
   "Z201".tInputs.xM209FanProtection :="FB_CommunicationZ300_V1.00_DB".IN_tIDeviceDataIN.Z200.IN_MCC1201."xA.E83.5";
   "Z201".tInputs.xM209FanFeedback := "FB_CommunicationZ300_V1.00_DB".IN_tIDeviceDataIN.Z200.IN_MCC1201."xA.E83.6";

   "FB_ManInsp_V1_00_IDB".INPUT.rgxQualityButtons[1]:="FB_CommunicationZ300_V1.00_DB".IN_tIDeviceDataIN.Z200.IN_MCC1301."xE.E108.4";


   "FB_DropConveyor_IDB".INPUT.xUpPosition := "FB_CommunicationZ300_V1.00_DB".IN_tIDeviceDataIN.Z200.IN_MCC1201."xA.E82.1";
   "FB_DropConveyor_IDB".INPUT.xDownPosition := "FB_CommunicationZ300_V1.00_DB".IN_tIDeviceDataIN.Z200.IN_MCC1201."xA.E82.2";
   "FB_DropConveyor_IDB".INPUT.xDoorOpen := "FB_CommunicationZ300_V1.00_DB".IN_tIDeviceDataIN.Z200.IN_MCC1201."xA.E34.0"OR"FB_CommunicationZ300_V1.00_DB".IN_tIDeviceDataIN.Z200.IN_MCC1201."xA.E34.7" ;
   "FB_DropConveyor_IDB".INPUT.xFeedbackMovement :="FB_CommunicationZ300_V1.00_DB".IN_tIDeviceDataIN.Z200.IN_MCC1201."xA.E82.0" ;
   "FB_DropConveyor_IDB".INPUT.xProtection :="FB_CommunicationZ300_V1.00_DB".IN_tIDeviceDataIN.Z200.IN_MCC1201."xA.E81.5" ;
   "FB_DropConveyor_IDB".INPUT.xProtectionBrake := 1;
   "FB_DropConveyor_IDB".INPUT.xUpDownPushbutton := "FB_CommunicationZ300_V1.00_DB".IN_tIDeviceDataIN.Z200.IN_MCC1201."xA.E35.0" OR"FB_CommunicationZ300_V1.00_DB".IN_tIDeviceDataIN.Z200.IN_MCC1201."xA.E34.2" ;
   "FB_DropConveyor_IDB".INPUT.xSafetyBar := "FB_CommunicationZ300_V1.00_DB".IN_tIDeviceDataIN.Z200.IN_MCC1201."xA.E82.3";

   "FB_BreakerM206_V1_00_IDB".INPUT.xConditionOKFromCulletSystem := "FB_CommunicationZ300_V1.00_DB".IN_tIDeviceDataIN.Z200.IN_MCC1201."xA.E39.0";
   "FB_BreakerM206_V1_00_IDB".INPUT.xBreakerRotationControl := "FB_CommunicationZ300_V1.00_DB".IN_tIDeviceDataIN.Z200.IN_MCC1201."xA.E36.0";
   "FB_BreakerM206_V1_00_IDB".INPUT.xProtectionBreakerRotation := "FB_CommunicationZ300_V1.00_DB".IN_tIDeviceDataIN.Z200.IN_MCC1201."xA.E83.0";
   "FB_BreakerM206_V1_00_IDB".INPUT.xFeedbackRotationKM := "FB_CommunicationZ300_V1.00_DB".IN_tIDeviceDataIN.Z200.IN_MCC1201."xA.E83.1";

   "FB_IO_EmergencyCuttingBridge_DB".IN_xMachineReady :="FB_CommunicationZ300_V1.00_DB".IN_tIDeviceDataIN.Z200.IN_MCC1201."xA.E33.4";
   "FB_IO_EmergencyCuttingBridge_DB".IN_xStartCutCycle := "FB_CommunicationZ300_V1.00_DB".IN_tIDeviceDataIN.Z200.IN_MCC1201."xA.E33.5";
   "FB_IO_EmergencyCuttingBridge_DB".IN_xProtection := "FB_CommunicationZ300_V1.00_DB".IN_tIDeviceDataIN.Z200.IN_MCC1201."xA.E81.2";

   "FB_BD_BreakPH_V1_00_IDB".INPUT.rgxPhotoStatus[0] := "FB_CommunicationZ300_V1.00_DB".IN_tIDeviceDataIN.Z200.IN_MCC1201."xA.E32.0";
   "FB_BD_BreakPH_V1_00_IDB".INPUT.rgxPhotoStatus[1]:= "FB_CommunicationZ300_V1.00_DB".IN_tIDeviceDataIN.Z200.IN_MCC1201."xA.E32.1";
   "FB_BD_BreakPH_V1_00_IDB".INPUT.rgxPhotoStatus[2] := "FB_CommunicationZ300_V1.00_DB".IN_tIDeviceDataIN.Z200.IN_MCC1201."xA.E32.2";
   "FB_BD_BreakPH_V1_00_IDB".INPUT.rgxPhotoStatus[3] := "FB_CommunicationZ300_V1.00_DB".IN_tIDeviceDataIN.Z200.IN_MCC1201."xA.E32.3";
   "FB_BD_BreakPH_V1_00_IDB".INPUT.rgxPhotoStatus[4] := "FB_CommunicationZ300_V1.00_DB".IN_tIDeviceDataIN.Z200.IN_MCC1201."xA.E32.4";
   "FB_BD_BreakPH_V1_00_IDB".INPUT.rgxPhotoStatus[5] := "FB_CommunicationZ300_V1.00_DB".IN_tIDeviceDataIN.Z200.IN_MCC1201."xA.E32.5";
   "FB_BD_BreakPH_V1_00_IDB".INPUT.rgxPhotoStatus[6] := "FB_CommunicationZ300_V1.00_DB".IN_tIDeviceDataIN.Z200.IN_MCC1201."xA.E32.6";
   "FB_BD_BreakPH_V1_00_IDB".INPUT.rgxPhotoStatus[7] := "FB_CommunicationZ300_V1.00_DB".IN_tIDeviceDataIN.Z200.IN_MCC1201."xA.E32.7";
   "FB_BD_BreakPH_V1_00_IDB".INPUT.rgxPhotoStatus[8] := "FB_CommunicationZ300_V1.00_DB".IN_tIDeviceDataIN.Z200.IN_MCC1201."xA.E33.0";
   "FB_BD_BreakPH_V1_00_IDB".INPUT.rgxPhotoStatus[9] := "FB_CommunicationZ300_V1.00_DB".IN_tIDeviceDataIN.Z200.IN_MCC1201."xA.E33.1";

   "FB_BD_BreakPH_V1_00_IDB".INPUT.xButtonAlarmOFF:="FB_CommunicationZ300_V1.00_DB".IN_tIDeviceDataIN.Z200.IN_MCC1301."xE.E108.6" OR"FB_CommunicationZ300_V1.00_DB".IN_tIDeviceDataIN.Z200.IN_MCC1201."xA.E34.1";

   "FB_Z200Conveyor_M201_IDB".INPUT_xLocalSwitch := TRUE;
   "FB_Z200Conveyor_M201_IDB".INPUT_xMotorThermalProbe := "FB_CommunicationZ300_V1.00_DB".IN_tIDeviceDataIN.Z200.IN_MCC1201."xA.E38.6";
   "FB_Z200Conveyor_M201_IDB".INPUT_xQFMotorFan := "CU_A250AP1_IDB".STC_tPZD_CU.tR.tE_DIGITAL.x9;
   "FB_Z200Conveyor_M201_IDB".INPUT_xPowerModuleOn := "CU_A250AP1_IDB".OUT_xPower_ON;
   //"FB_Z200Conveyor_M201_IDB".INPUT_dMagnitude := "IN_dMagnitude_M201";
   //"FB_Z200Conveyor_M201_IDB".INPUT_dTorque := "IN_dTorque_M201";


   "FB_Z200Conveyor_M204_IDB".INPUT_xLocalSwitch := TRUE;
   "FB_Z200Conveyor_M204_IDB".INPUT_xMotorThermalProbe := "FB_CommunicationZ300_V1.00_DB".IN_tIDeviceDataIN.Z200.IN_MCC1201."xA.E38.7";
   "FB_Z200Conveyor_M204_IDB".INPUT_xQFMotorFan := "CU_A250AP1_IDB".STC_tPZD_CU.tR.tE_DIGITAL.x10;
   "FB_Z200Conveyor_M204_IDB".INPUT_xPowerModuleOn := "CU_A250AP1_IDB".OUT_xPower_ON;
   //"FB_Z200Conveyor_M204_IDB".INPUT_dMagnitude := "IN_dMagnitude_M204";
   //"FB_Z200Conveyor_M204_IDB".INPUT_dTorque := "IN_dTorque_M204";


   "FB_Z200Conveyor_M205_IDB".INPUT_xLocalSwitch := TRUE;
   "FB_Z200Conveyor_M205_IDB".INPUT_xMotorThermalProbe := "FB_CommunicationZ300_V1.00_DB".IN_tIDeviceDataIN.Z200.IN_MCC1201."xA.E39.3";
   "FB_Z200Conveyor_M205_IDB".INPUT_xQFMotorFan :=TRUE;
   "FB_Z200Conveyor_M205_IDB".INPUT_xPowerModuleOn := "CU_A260AP1_IDB".OUT_xPower_ON;
   //"FB_Z200Conveyor_M205_IDB".INPUT_dMagnitude := "IN_dMagnitude_M208";
   //"FB_Z200Conveyor_M205_IDB".INPUT_dTorque := "IN_dTorque_M208";

   "FB_Z200Conveyor_M208_IDB".INPUT_xLocalSwitch := TRUE;
   "FB_Z200Conveyor_M208_IDB".INPUT_xMotorThermalProbe := "FB_CommunicationZ300_V1.00_DB".IN_tIDeviceDataIN.Z200.IN_MCC1201."xA.E39.4";
   "FB_Z200Conveyor_M208_IDB".INPUT_xQFMotorFan :=  "CU_A260AP1_IDB".STC_tPZD_CU.tR.tE_DIGITAL.x9;
   "FB_Z200Conveyor_M208_IDB".INPUT_xPowerModuleOn := "CU_A260AP1_IDB".OUT_xPower_ON;
   //"FB_Z200Conveyor_M208_IDB".INPUT_dMagnitude := "IN_dMagnitude_M208";
   //"FB_Z200Conveyor_M208_IDB".INPUT_dTorque := "IN_dTorque_M208";

   "FB_Z200Conveyor_M211_iDB".INPUT_xLocalSwitch := TRUE;
   "FB_Z200Conveyor_M211_iDB".INPUT_xMotorThermalProbe := "FB_CommunicationZ300_V1.00_DB".IN_tIDeviceDataIN.Z200.IN_MCC1201."xA.E39.5";
   "FB_Z200Conveyor_M211_iDB".INPUT_xQFMotorFan := "CU_A260AP1_IDB".STC_tPZD_CU.tR.tE_DIGITAL.x10;
   "FB_Z200Conveyor_M211_iDB".INPUT_xPowerModuleOn := "CU_A260AP1_IDB".OUT_xPower_ON;
   //"FB_Z200Conveyor_M211_IDB".INPUT_dMagnitude := "IN_dMagnitude_M211";
   //"FB_Z200Conveyor_M211_IDB".INPUT_dTorque := "IN_dTorque_M211";

   "FB_Z200Conveyor_M214_iDB".INPUT_xLocalSwitch := TRUE;
   "FB_Z200Conveyor_M214_iDB".INPUT_xMotorThermalProbe := "FB_CommunicationZ300_V1.00_DB".IN_tIDeviceDataIN.Z200.IN_MCC1201."xA.E39.6";
   "FB_Z200Conveyor_M214_iDB".INPUT_xQFMotorFan := "CU_A260AP1_IDB".STC_tPZD_CU.tR.tE_DIGITAL.x11;
   "FB_Z200Conveyor_M214_iDB".INPUT_xPowerModuleOn := "CU_A260AP1_IDB".OUT_xPower_ON;
   //"FB_Z200Conveyor_M214_IDB".INPUT_dMagnitude := "IN_dMagnitude_M214";
   //"FB_Z200Conveyor_M214_IDB".INPUT_dTorque := "IN_dTorque_M214";


   "FB_Z200Conveyor_M218_IDB".INPUT_xLocalSwitch := TRUE;
   "FB_Z200Conveyor_M218_IDB".INPUT_xMotorThermalProbe := "FB_CommunicationZ300_V1.00_DB".IN_tIDeviceDataIN.Z200.IN_MCC1201."xA.E39.7";
   "FB_Z200Conveyor_M218_IDB".INPUT_xQFMotorFan := "CU_A260AP1_IDB".STC_tPZD_CU.tR.tE_DIGITAL_1.x8;
   "FB_Z200Conveyor_M218_IDB".INPUT_xPowerModuleOn := "CU_A260AP1_IDB".OUT_xPower_ON;
   //"FB_Z200Conveyor_M218_IDB".INPUT_dMagnitude := "IN_dMagnitude_M218";
   //"FB_Z200Conveyor_M218_IDB".INPUT_dTorque := "IN_dTorque_M218";

   "DB_AUX_Z200_SpeedLehr".dPulseEncoder1 := "FB_CommunicationZ300_V1.00_DB".IN_tIDeviceDataIN.Z200.dLherSpeed_Enc1;
   "DB_AUX_Z200_SpeedLehr".dPulseEncoder2 := "FB_CommunicationZ300_V1.00_DB".IN_tIDeviceDataIN.Z200.dLherSpeed_Enc2;
END_REGION
END_FUNCTION

// folder: 03_Programs_Logics/MCC1200/01_Defects

FUNCTION_BLOCK "FB_TrackDefects_V1.00"   // FB16, LAD
TITLE = Tracking defects
{ S7_Optimized_Access := 'TRUE' }
VERSION : 0.1
   VAR_INPUT
      IN_xFaultsEnabled : Bool;   // Faults enabled
      IN_xCycleON : Bool;   // Zone is in cycle
      IN_xGeneralReset : Bool;   // General reset
      IN_xFaultsReset : Bool;   // Reset alarms
      IN_xSimulationActive : Bool;   // Simulation active
      IN_dSimSendRate_ms : DInt;   // Simulation defect sending rate [ms]
      IN_dSimMaxClass : DInt;   // Simulation max class
      IN_dSimMinYPos_cmm : DInt;   // Simulation minimum Y position [mm/100]
      IN_dSimMaxYPos_cmm : DInt;   // Simulation maximum Y position [mm/100]
      IN_dSimXPosInsert_cmm : DInt;   // Simulation position X [mm/100]
   END_VAR
   VAR_IN_OUT
      INO_tEncoder : "UDT_Encoder";   // Encoder data
      INO_tDefects : "UDT_DefectData_Tracking_Ext";   // Defects data
      INO_tOBInit : "GP_OB_Initialize";
      INO_tFBAddSlow : "FB_Defects_Add_V1.00";   // Defect tank slow task
      INO_tFBAddMed : "FB_Defects_Add_V1.00";   // Defect tank medium task
      INO_tFBAddFast : "FB_Defects_Add_V1.00";   // Defect tank fast task
      INO_tFBAddMain : "FB_Defects_Add_V1.00";   // Defect tank main task
   END_VAR
   VAR
      OSR_xGeneralReset : Bool;   // OSR.General reset
      AUX_tEmptyDefect : "UDT_DefectDataExt";   // Always empty defect
      AUX_dSimLastGenDef : DInt;   // Simulation last generated defect
      AUX_dtActDate : DTL;
   END_VAR
   VAR_TEMP
      TMP_xOSGeneralReset : Bool;
      TMP_dIndex : DInt;
      TMP_dValue_cmm : DInt;
      TMP_dNextTail : DInt;
      TMP_dNextHead : DInt;
      TMP_xRandOut : Bool;
      TMP_uiRandStatus : UInt;
      TMP_wStatus : Word;
      TMP_dClass : DInt;
      TMP_dDefYPos_cmm : DInt;
      TMP_dDefXPos_cmm : DInt;
      TMP_iDummy : Int;
      TMP_strDateTime : String;
   END_VAR
   VAR CONSTANT
      CONST_DTHRDELDEFECT_CMM : DInt := 200000;   // Threshold delete defect [mm/100]
      CONST_DMAXIDDEFECTS : DInt := 2000000000;   // Maximum defect ID
   END_VAR
   VAR_TEMP   // added for the SCL form of the ladder/FBD networks
      _w1 : Bool;
   END_VAR
BEGIN

REGION Network 1: General reset
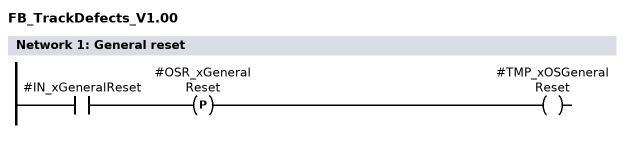
   RUNG wire#powerrail
      Contact( #IN_xGeneralReset )
      P_Trig( #OSR_xGeneralReset )
      Coil( #TMP_xOSGeneralReset )
   END_RUNG
   // the same network as SCL:
   #_w1 := #IN_xGeneralReset AND NOT #OSR_xGeneralReset;   // rising edge
   #OSR_xGeneralReset := #IN_xGeneralReset;
   #TMP_xOSGeneralReset := #_w1;
END_REGION

REGION Network 2 (SCL): Reset all the buffers
   IF #TMP_xOSGeneralReset THEN

       #INO_tDefects.dBufferHead := -1;
       #INO_tDefects.dBufferTail := -1;
       #INO_tDefects.dBufferTailOptimizer := -1;
       #INO_tDefects.dBufferTailReport := -1;
       #INO_tDefects.dBufferTailOptPLC := -1;
       #INO_tDefects.tDefectsForOpt.dNumberOfDefect := 0;
       #INO_tDefects.tDefectsForReport.dNumberOfDefect := 0;    
       #INO_tDefects.tDefectsforOptPlc.dNumberOfDefect := 0;    

       FOR #TMP_dIndex := 0 TO "DNUMDEFFOROPT_IND" DO
           #INO_tDefects.tDefectsForOpt.rgtDefects[#TMP_dIndex] := #AUX_tEmptyDefect;
       END_FOR;

       FOR #TMP_dIndex := 0 TO "DNUMDEFFOROPT_IND" DO
           #INO_tDefects.tDefectsforOptPlc.rgtDefects[#TMP_dIndex] := #AUX_tEmptyDefect;
       END_FOR;

       FOR #TMP_dIndex := 0 TO "DNUMDEFFORREPORT_IND" DO
           #INO_tDefects.tDefectsForReport.rgtDefects[#TMP_dIndex] := #AUX_tEmptyDefect;
       END_FOR;

       FOR #TMP_dIndex := 0 TO "DNUMDEFEXT_IND" DO

           #INO_tDefects.rgtDefects[#TMP_dIndex] := #AUX_tEmptyDefect;

       END_FOR;

   END_IF;
END_REGION

REGION Network 3 (SCL): Delete defect on buffer
   //At the moment this delete is disabled, is better keep all the defect in case of optimizer need.
   (*
   WHILE   (#INO_tDefects.dBufferTail <> #INO_tDefects.dBufferHead) AND
           (#INO_tDefects.dBufferTail <> #INO_tDefects.dBufferTailOptimizer) AND
           (#INO_tDefects.dBufferTailReport = #INO_tDefects.dBufferTailOptimizer) DO

       #INO_tDefects.rgtDefects[#INO_tDefects.dBufferTail] := #AUX_tEmptyDefect;

       IF (#INO_tDefects.dBufferTail + 1) >= "DNUMDEFEXT" THEN
           #INO_tDefects.dBufferTail := 0;
       ELSE
           #INO_tDefects.dBufferTail := #INO_tDefects.dBufferTail + 1;
       END_IF;

   END_WHILE;
   *)
END_REGION

REGION Network 4 (SCL): Delete defect on buffer after position
   WHILE (#INO_tDefects.dBufferTail <> #INO_tDefects.dBufferHead) AND (#INO_tDefects.dBufferHead <> -1) DO

       IF (#INO_tDefects.dBufferTail + 1) >= "DNUMDEFEXT" THEN
           #TMP_dNextTail := 0;
       ELSE
           #TMP_dNextTail := #INO_tDefects.dBufferTail + 1;
       END_IF;

       #TMP_dValue_cmm := #INO_tEncoder.dActualEncoderCounter_cmm - #INO_tDefects.rgtDefects[#TMP_dNextTail].dXPosition_cmm;

       IF (#TMP_dValue_cmm > #CONST_DTHRDELDEFECT_CMM) THEN

           #INO_tDefects.rgtDefects[#TMP_dNextTail] := #AUX_tEmptyDefect;

           IF (#INO_tDefects.dBufferTail = #INO_tDefects.dBufferTailOptPLC) THEN
               #INO_tDefects.dBufferTailOptPLC := #TMP_dNextTail;
           END_IF;

           IF (#INO_tDefects.dBufferTail = #INO_tDefects.dBufferTailOptimizer) THEN
               #INO_tDefects.dBufferTailOptimizer := #TMP_dNextTail;
           END_IF;

           IF (#INO_tDefects.dBufferTail = #INO_tDefects.dBufferTailReport) THEN
               #INO_tDefects.dBufferTailReport := #TMP_dNextTail;
           END_IF;

           #INO_tDefects.dBufferTail := #TMP_dNextTail;

       ELSE
           EXIT; //Exit the while
       END_IF;    

   END_WHILE;
END_REGION

REGION Network 5 (SCL): Insert defect from buffer slow
   IF (#INO_tFBAddSlow.ST_xDefectIsUpdating = FALSE) AND (#INO_tFBAddSlow.AUX_dNumDefectOnBuffer > 0) THEN

       #TMP_dIndex := #INO_tFBAddSlow.AUX_dNumDefectOnBuffer - 1;

       WHILE (#TMP_dIndex >= 0) DO

           //Increment the index head
           IF (#INO_tDefects.dBufferHead + 1) >= "DNUMDEFEXT" THEN
               #TMP_dNextHead := 0;
           ELSE
               #TMP_dNextHead := #INO_tDefects.dBufferHead + 1;
           END_IF;

           //Check if the buffer is full
           IF (#TMP_dNextHead = #INO_tDefects.dBufferTail) AND (#INO_tDefects.dBufferHead <> -1) THEN
               EXIT;
           END_IF; 

           #INO_tDefects.rgtDefects[#TMP_dNextHead] := #INO_tFBAddSlow.AUX_rgtDefects[#TMP_dIndex];
           #INO_tDefects.rgtDefects[#TMP_dNextHead].dID := #INO_tDefects.dDefectNextID;

           //Reset to 0 the data
           //#INO_tFBAddSlow.AUX_rgtDefects[#TMP_dIndex] := #AUX_tEmptyDefect;

           #TMP_dIndex -= 1;
           #INO_tFBAddSlow.AUX_dNumDefectOnBuffer -= 1;
           #INO_tDefects.dBufferHead := #TMP_dNextHead;

           #INO_tDefects.dDefectNextID += 1;

           IF #INO_tDefects.dDefectNextID > #CONST_DMAXIDDEFECTS THEN
               #INO_tDefects.dDefectNextID := 1;
           END_IF;

       END_WHILE;
   END_IF;
END_REGION

REGION Network 6 (SCL): Insert defect from buffer medium
   IF (#INO_tFBAddMed.ST_xDefectIsUpdating = FALSE) AND (#INO_tFBAddMed.AUX_dNumDefectOnBuffer > 0) THEN

       #TMP_dIndex := #INO_tFBAddMed.AUX_dNumDefectOnBuffer - 1;

       WHILE (#TMP_dIndex >= 0) DO

           //Increment the index head
           IF (#INO_tDefects.dBufferHead + 1) >= "DNUMDEFEXT" THEN
               #TMP_dNextHead := 0;
           ELSE
               #TMP_dNextHead := #INO_tDefects.dBufferHead + 1;
           END_IF;

           //Check if the buffer is full
           IF (#TMP_dNextHead = #INO_tDefects.dBufferTail) AND (#INO_tDefects.dBufferHead <> -1) THEN
               EXIT;
           END_IF; 

           #INO_tDefects.rgtDefects[#TMP_dNextHead] := #INO_tFBAddMed.AUX_rgtDefects[#TMP_dIndex];
           #INO_tDefects.rgtDefects[#TMP_dNextHead].dID := #INO_tDefects.dDefectNextID;

           //Reset to 0 the data
           #INO_tFBAddMed.AUX_rgtDefects[#TMP_dIndex] := #AUX_tEmptyDefect;

           #TMP_dIndex -= 1;
           #INO_tFBAddMed.AUX_dNumDefectOnBuffer -= 1;
           #INO_tDefects.dBufferHead := #TMP_dNextHead;

           #INO_tDefects.dDefectNextID += 1;

           IF #INO_tDefects.dDefectNextID > #CONST_DMAXIDDEFECTS THEN
               #INO_tDefects.dDefectNextID := 1;
           END_IF;

       END_WHILE;

   END_IF;
END_REGION

REGION Network 7 (SCL): Insert defect from buffer fast
   IF (#INO_tFBAddFast.ST_xDefectIsUpdating = FALSE) AND (#INO_tFBAddFast.AUX_dNumDefectOnBuffer > 0) THEN

       #TMP_dIndex := #INO_tFBAddFast.AUX_dNumDefectOnBuffer - 1;

       WHILE (#TMP_dIndex >= 0) DO

           //Increment the index head
           IF (#INO_tDefects.dBufferHead + 1) >= "DNUMDEFEXT" THEN
               #TMP_dNextHead := 0;
           ELSE
               #TMP_dNextHead := #INO_tDefects.dBufferHead + 1;
           END_IF;

           //Check if the buffer is full
           IF (#TMP_dNextHead = #INO_tDefects.dBufferTail) AND (#INO_tDefects.dBufferHead <> -1) THEN
               EXIT;
           END_IF; 

           #INO_tDefects.rgtDefects[#TMP_dNextHead] := #INO_tFBAddFast.AUX_rgtDefects[#TMP_dIndex];
           #INO_tDefects.rgtDefects[#TMP_dNextHead].dID := #INO_tDefects.dDefectNextID;

           //Reset to 0 the data
           #INO_tFBAddFast.AUX_rgtDefects[#TMP_dIndex] := #AUX_tEmptyDefect;

           #TMP_dIndex -= 1;
           #INO_tFBAddFast.AUX_dNumDefectOnBuffer -= 1;
           #INO_tDefects.dBufferHead := #TMP_dNextHead;

           #INO_tDefects.dDefectNextID += 1;

           IF #INO_tDefects.dDefectNextID > #CONST_DMAXIDDEFECTS THEN
               #INO_tDefects.dDefectNextID := 1;
           END_IF;

       END_WHILE;

   END_IF;
END_REGION

REGION Network 8 (SCL): Insert defect from buffer main
   IF (#INO_tFBAddMain.ST_xDefectIsUpdating = FALSE) AND (#INO_tFBAddMain.AUX_dNumDefectOnBuffer > 0) THEN

       #TMP_dIndex := #INO_tFBAddMain.AUX_dNumDefectOnBuffer - 1;

       WHILE (#TMP_dIndex >= 0) DO

           //Increment the index head
           IF (#INO_tDefects.dBufferHead + 1) >= "DNUMDEFEXT" THEN
               #TMP_dNextHead := 0;
           ELSE
               #TMP_dNextHead := #INO_tDefects.dBufferHead + 1;
           END_IF;

           //Check if the buffer is full
           IF (#TMP_dNextHead = #INO_tDefects.dBufferTail)AND (#INO_tDefects.dBufferHead <> -1) THEN
               EXIT;
           END_IF; 

           #INO_tDefects.rgtDefects[#TMP_dNextHead] := #INO_tFBAddMain.AUX_rgtDefects[#TMP_dIndex];
           #INO_tDefects.rgtDefects[#TMP_dNextHead].dID := #INO_tDefects.dDefectNextID;

           //Reset to 0 the data
           #INO_tFBAddMain.AUX_rgtDefects[#TMP_dIndex] := #AUX_tEmptyDefect;

           #TMP_dIndex -= 1;
           #INO_tFBAddMain.AUX_dNumDefectOnBuffer -= 1;
           #INO_tDefects.dBufferHead := #TMP_dNextHead;

           #INO_tDefects.dDefectNextID += 1;

           IF #INO_tDefects.dDefectNextID > #CONST_DMAXIDDEFECTS THEN
               #INO_tDefects.dDefectNextID := 1;
           END_IF;

       END_WHILE;

   END_IF;
END_REGION

REGION Network 9 (SCL): Prepare defect for report
   IF (#INO_tDefects.tDefectsForReport.dNumberOfDefect = 0)  THEN

       #TMP_dIndex := 0;

       WHILE ((#TMP_dIndex <= "DNUMDEFFORREPORT_IND") AND (#INO_tDefects.dBufferTailReport <> #INO_tDefects.dBufferHead) AND  (#INO_tDefects.dBufferHead <> -1)) DO

           IF (#INO_tDefects.dBufferTailReport + 1) >= "DNUMDEFEXT" THEN
               #TMP_dNextTail := 0;
           ELSE
               #TMP_dNextTail := #INO_tDefects.dBufferTailReport + 1;
           END_IF;

           #INO_tDefects.tDefectsForReport.rgtDefects[#TMP_dIndex] := #INO_tDefects.rgtDefects[#TMP_dNextTail];

           #INO_tDefects.dBufferTailReport := #TMP_dNextTail;

           #TMP_dIndex += 1;

       END_WHILE;

       #INO_tDefects.tDefectsForReport.dNumberOfDefect := #TMP_dIndex;

       IF #INO_tDefects.tDefectsForReport.dNumberOfDefect > 0 THEN    
           FOR #TMP_dIndex := #INO_tDefects.tDefectsForReport.dNumberOfDefect TO "DNUMDEFFORREPORT_IND" DO
               #INO_tDefects.tDefectsForReport.rgtDefects[#TMP_dIndex] := #AUX_tEmptyDefect;
           END_FOR;
       END_IF;

   ELSE
       //Check the first defects, if is too old delete the whole buffer
      #TMP_dValue_cmm := #INO_tEncoder.dActualEncoderCounter_cmm - #INO_tDefects.tDefectsForReport.rgtDefects[0].dXPosition_cmm;

       IF (#TMP_dValue_cmm > (#CONST_DTHRDELDEFECT_CMM * 10)) THEN

           FOR #TMP_dIndex := 0 TO #INO_tDefects.tDefectsForReport.dNumberOfDefect - 1 DO

               #INO_tDefects.tDefectsForReport.rgtDefects[#TMP_dIndex] := #AUX_tEmptyDefect;

           END_FOR;

           #INO_tDefects.tDefectsForReport.dNumberOfDefect := 0;

       END_IF;

   END_IF;
END_REGION

REGION Network 10 (SCL): BPS / OPTs require to resend all defects
   IF #INO_tDefects.xBPSARequireAllDef THEN
       #INO_tDefects.xBPSARequireAllDef := FALSE;
       #INO_tDefects.dBufferTailReport := #INO_tDefects.dBufferTail;    
   END_IF;

   IF #INO_tDefects.xBPSBRequireAllDef THEN
       #INO_tDefects.xBPSBRequireAllDef := FALSE;
       #INO_tDefects.dBufferTailReport := #INO_tDefects.dBufferTail;    
   END_IF;

   IF #INO_tDefects.xOptimizerRequireAllDef THEN
       #INO_tDefects.xOptimizerRequireAllDef := FALSE;
       #INO_tDefects.dBufferTailOptimizer := #INO_tDefects.dBufferTail;    

   END_IF;

   IF #INO_tDefects.xOptimizerPLCRequireAllDef THEN
       #INO_tDefects.xOptimizerPLCRequireAllDef := FALSE;
       #INO_tDefects.dBufferTailOptPLC := #INO_tDefects.dBufferTail;    
   END_IF;
END_REGION

REGION Network 11 (SCL): Prepare defect for optimizer
   IF (#INO_tDefects.tDefectsForOpt.dNumberOfDefect = 0) AND (#INO_tDefects.dBufferHead <> -1)THEN

       #TMP_dIndex := 0;

       WHILE ((#TMP_dIndex <= "DNUMDEFFOROPT_IND") AND (#INO_tDefects.dBufferTailOptimizer <> #INO_tDefects.dBufferHead) AND  (#INO_tDefects.dBufferHead <> -1)) DO

           IF (#INO_tDefects.dBufferTailOptimizer + 1) >= "DNUMDEFEXT" THEN
               #TMP_dNextTail := 0;
           ELSE
               #TMP_dNextTail := #INO_tDefects.dBufferTailOptimizer + 1;
           END_IF;

           #INO_tDefects.tDefectsForOpt.rgtDefects[#TMP_dIndex] := #INO_tDefects.rgtDefects[#TMP_dNextTail];

           #INO_tDefects.dBufferTailOptimizer := #TMP_dNextTail;

           #TMP_dIndex += 1;

       END_WHILE;

       #INO_tDefects.tDefectsForOpt.dNumberOfDefect := #TMP_dIndex;

       FOR #TMP_dIndex := #INO_tDefects.tDefectsForOpt.dNumberOfDefect TO "DNUMDEFFOROPT_IND" DO
           #INO_tDefects.tDefectsForOpt.rgtDefects[#TMP_dIndex] := #AUX_tEmptyDefect;
       END_FOR;

   ELSE
       //Check the first defects, if is too old delete the whole buffer
       #TMP_dValue_cmm := #INO_tEncoder.dActualEncoderCounter_cmm - #INO_tDefects.tDefectsForOpt.rgtDefects[0].dXPosition_cmm;

       IF (#TMP_dValue_cmm > (#CONST_DTHRDELDEFECT_CMM * 10)) THEN

           FOR #TMP_dIndex := 0 TO #INO_tDefects.tDefectsForOpt.dNumberOfDefect - 1 DO

               #INO_tDefects.tDefectsForOpt.rgtDefects[#TMP_dIndex] := #AUX_tEmptyDefect;

           END_FOR;

           #INO_tDefects.tDefectsForOpt.dNumberOfDefect := 0;

       END_IF;
   END_IF;
END_REGION

REGION Network 12 (SCL): Prepare defect for optimizer PLC
   IF (#INO_tDefects.tDefectsforOptPlc.dNumberOfDefect = 0) AND (#INO_tDefects.dBufferHead <> -1)THEN

       #TMP_dIndex := 0;

       WHILE ((#TMP_dIndex <= "DNUMDEFFOROPT_IND") AND (#INO_tDefects.dBufferTailOptPLC <> #INO_tDefects.dBufferHead) AND  (#INO_tDefects.dBufferHead <> -1)) DO

           IF (#INO_tDefects.dBufferTailOptPLC + 1) >= "DNUMDEFEXT" THEN
               #TMP_dNextTail := 0;
           ELSE
               #TMP_dNextTail := #INO_tDefects.dBufferTailOptPLC + 1;
           END_IF;

           #INO_tDefects.tDefectsforOptPlc.rgtDefects[#TMP_dIndex] := #INO_tDefects.rgtDefects[#TMP_dNextTail];

           #INO_tDefects.dBufferTailOptPLC := #TMP_dNextTail;

           #TMP_dIndex += 1;

       END_WHILE;

       #INO_tDefects.tDefectsforOptPlc.dNumberOfDefect := #TMP_dIndex;

       FOR #TMP_dIndex := #INO_tDefects.tDefectsforOptPlc.dNumberOfDefect TO "DNUMDEFFOROPT_IND" DO
           #INO_tDefects.tDefectsforOptPlc.rgtDefects[#TMP_dIndex] := #AUX_tEmptyDefect;
       END_FOR;

   ELSE
       //Check the first defects, if is too old delete the whole buffer
       #TMP_dValue_cmm := #INO_tEncoder.dActualEncoderCounter_cmm - #INO_tDefects.tDefectsforOptPlc.rgtDefects[0].dXPosition_cmm;

       IF (#TMP_dValue_cmm > (#CONST_DTHRDELDEFECT_CMM * 10)) THEN

           FOR #TMP_dIndex := 0 TO #INO_tDefects.tDefectsforOptPlc.dNumberOfDefect - 1 DO

               #INO_tDefects.tDefectsforOptPlc.rgtDefects[#TMP_dIndex] := #AUX_tEmptyDefect;

           END_FOR;

           #INO_tDefects.tDefectsforOptPlc.dNumberOfDefect := 0;

       END_IF;
   END_IF;
END_REGION

REGION Network 14 (SCL): ### SIMULATION ###
   #AUX_dSimLastGenDef -= #INO_tOBInit.OUT_dExecutionTime_ms;

   IF #AUX_dSimLastGenDef < 0 THEN
       #AUX_dSimLastGenDef := 0;
   END_IF;

   IF (#IN_xSimulationActive) AND (#AUX_dSimLastGenDef <= 0) THEN

       #AUX_dSimLastGenDef := #IN_dSimSendRate_ms;

       #TMP_dClass := "LGF_RandomRange_Dint"(minValue:=1, maxValue:=DINT_TO_INT(#IN_dSimMaxClass), error=>#TMP_xRandOut, subfunctionStatus=>#TMP_wStatus, status=>#TMP_wStatus);
       #TMP_dDefYPos_cmm := REAL_TO_DINT("LGF_RandomRange_Real"(minValue:=DINT_TO_REAL(#IN_dSimMinYPos_cmm), maxValue:=DINT_TO_REAL(#IN_dSimMaxYPos_cmm), error=>#TMP_xRandOut, subfunctionStatus=>#TMP_uiRandStatus, status=>#TMP_wStatus));
       #TMP_dDefXPos_cmm := #INO_tEncoder.dActualEncoderCounter_cmm + #IN_dSimXPosInsert_cmm;

       //Increment the index head
       IF (#INO_tDefects.dBufferHead + 1) >= "DNUMDEFEXT" THEN
           #TMP_dNextHead := 0;
       ELSE
           #TMP_dNextHead := #INO_tDefects.dBufferHead + 1;
       END_IF;

       //Check if the buffer is full
       IF (#TMP_dNextHead <> #INO_tDefects.dBufferTail) OR (#INO_tDefects.dBufferHead = -1) THEN

           #INO_tDefects.rgtDefects[#TMP_dNextHead].dID := #INO_tDefects.dDefectNextID;
           #INO_tDefects.rgtDefects[#TMP_dNextHead].dClass := #TMP_dClass;
           #INO_tDefects.rgtDefects[#TMP_dNextHead].dCoreLength_um := 1000;
           #INO_tDefects.rgtDefects[#TMP_dNextHead].dCoreWidth_um := 1000;
           #INO_tDefects.rgtDefects[#TMP_dNextHead].dDistLength_um := 2000;
           #INO_tDefects.rgtDefects[#TMP_dNextHead].dDistWidth_um := 2000;
           #INO_tDefects.rgtDefects[#TMP_dNextHead].dOptValue_mdptr := 0;
           #INO_tDefects.rgtDefects[#TMP_dNextHead].dSubType := 1;
           #INO_tDefects.rgtDefects[#TMP_dNextHead].dTotalLength_um := 3000;
           #INO_tDefects.rgtDefects[#TMP_dNextHead].dTotalWidth_um := 3000;
           #INO_tDefects.rgtDefects[#TMP_dNextHead].dXPosition_cmm := #TMP_dDefXPos_cmm;
           #INO_tDefects.rgtDefects[#TMP_dNextHead].dYPosition_cmm := #TMP_dDefYPos_cmm;

           #TMP_iDummy := RD_SYS_T(#AUX_dtActDate);

           #TMP_strDateTime := "LGF_DTLtoString_ISO"("date"  :=#AUX_dtActDate, separator:='-');

           #TMP_strDateTime := CONCAT(IN1:=#TMP_strDateTime, IN2:='#');
           #TMP_strDateTime := CONCAT(IN1:=#TMP_strDateTime, IN2:=DINT_TO_STRING(#INO_tDefects.dDefectNextID));

           #INO_tDefects.rgtDefects[#TMP_dNextHead].strDefectID := #TMP_strDateTime;


           #INO_tDefects.dBufferHead := #TMP_dNextHead;
           #INO_tDefects.dDefectNextID += 1;

           IF #INO_tDefects.dDefectNextID > #CONST_DMAXIDDEFECTS THEN
               #INO_tDefects.dDefectNextID := 1;
           END_IF;

       END_IF; 
   END_IF;
END_REGION
END_FUNCTION_BLOCK

FUNCTION_BLOCK "FB_Defects_Add_V1.00"   // FB17, LAD
{ S7_Optimized_Access := 'TRUE' }
VERSION : 0.1
   VAR_INPUT
      IN_dClass : DInt;   // Defect class value [Num]
      IN_dSubType : DInt;   // Defect subtype [Num]
      IN_dXPosition_cmm : DInt;   // Defect X position [mm/100]
      IN_dYPosition_cmm : DInt;   // Defect Y position [mm/100]
      IN_dTotalLength_um : DInt;   // Defect total length [um]
      IN_dTotalWidth_um : DInt;   // Defect total width [um]
      IN_dCoreLength_um : DInt;   // Defect core length [um]
      IN_dCoreWidth_um : DInt;   // Defect core width [um]
      IN_dDistLength_um : DInt;   // Defect distortion length [um]
      IN_dDistWidth_um : DInt;   // Defect distortion width [um]
      IN_dOptValue_mdptr : DInt;   // Defect optical distortion [mdptr]
      IN_strDefectID : String["DSTRSIZEDEFID"];   // Defect string ID
   END_VAR
   VAR_OUTPUT
      OUT_xBufferFull : Bool;   // Buffer is full (Retry to load the defect)
   END_VAR
   VAR
      AUX_dNumDefectOnBuffer : DInt;   // Number of defect on buffer
      AUX_rgtDefects : Array[0..#CONST_DMAXDEF_IND] of "UDT_DefectDataExt";   // Defect buffer
      ST_xDefectIsUpdating : Bool;   // Updating defect buffer (No read available)
   END_VAR
   VAR CONSTANT
      CONST_DMAXDEF : DInt := 50;   // Maximum number of defect on buffer
      CONST_DMAXDEF_IND : DInt := 49;   // Maximum number of defect on buffer -1 for index
   END_VAR
BEGIN

REGION Network 1 (SCL): Insert defect on the temporary buffer
   #ST_xDefectIsUpdating := TRUE;

   IF #AUX_dNumDefectOnBuffer < #CONST_DMAXDEF_IND THEN

       #OUT_xBufferFull := FALSE;

       #AUX_rgtDefects[#AUX_dNumDefectOnBuffer].dID := 0;
       #AUX_rgtDefects[#AUX_dNumDefectOnBuffer].dClass := #IN_dClass; 
       #AUX_rgtDefects[#AUX_dNumDefectOnBuffer].dSubType :=  #IN_dSubType;
       #AUX_rgtDefects[#AUX_dNumDefectOnBuffer].dXPosition_cmm := #IN_dXPosition_cmm;
       #AUX_rgtDefects[#AUX_dNumDefectOnBuffer].dYPosition_cmm := #IN_dYPosition_cmm; 
       #AUX_rgtDefects[#AUX_dNumDefectOnBuffer].dTotalLength_um := #IN_dTotalLength_um;  
       #AUX_rgtDefects[#AUX_dNumDefectOnBuffer].dTotalWidth_um := #IN_dTotalWidth_um;
       #AUX_rgtDefects[#AUX_dNumDefectOnBuffer].dCoreLength_um := #IN_dCoreLength_um;
       #AUX_rgtDefects[#AUX_dNumDefectOnBuffer].dCoreWidth_um := #IN_dCoreWidth_um;
       #AUX_rgtDefects[#AUX_dNumDefectOnBuffer].dDistLength_um := #IN_dDistLength_um;
       #AUX_rgtDefects[#AUX_dNumDefectOnBuffer].dDistWidth_um := #IN_dDistWidth_um;
       #AUX_rgtDefects[#AUX_dNumDefectOnBuffer].dOptValue_mdptr := #IN_dOptValue_mdptr;
       #AUX_rgtDefects[#AUX_dNumDefectOnBuffer].strDefectID :=  #IN_strDefectID;

       #AUX_dNumDefectOnBuffer += 1;

   ELSE
       #OUT_xBufferFull := TRUE;
   END_IF;

   #ST_xDefectIsUpdating := FALSE;
END_REGION
END_FUNCTION_BLOCK

// folder: 03_Programs_Logics/MCC1200/02_Plates

FUNCTION_BLOCK "FB_TrackCaps_V1.00"   // FB5, LAD
TITLE = Tracking caps
{ S7_Optimized_Access := 'TRUE' }
VERSION : 0.1
   VAR_INPUT
      IN_xFaultsEnabled : Bool;   // Faults enabled
      IN_xCycleON : Bool;   // Zone is in cycle
      IN_xGeneralReset : Bool;   // General reset
      IN_xFaultsReset : Bool;   // Reset alarms
   END_VAR
   VAR_IN_OUT
      INO_tCaps : "UDT_CapData_Tracking";   // Cap tracking
      INO_tEncoder : "UDT_Encoder";   // Encoder data
      INO_tOptManager : "FB_OptManager_V1.00";   // Optimizer manager
   END_VAR
   VAR
      STC_OSR_xGeneralReset : Bool;
   END_VAR
   VAR_TEMP
      TMP_dIndex : DInt;
      TMP_wValue : Word;
      TMP_dwValue : DWord;
      TMP_xOSGeneralReset : Bool;
      TMP_dValue_cmm : DInt;
      TMP_dActMachineEncValue_cmm : DInt;
      TMP_dIndexCap : DInt;
      TMP_xPlateFound : Bool;
      TMP_dTail : DInt;
      TMP_dHeadPosFromSnap_cmm : DInt;
      TMP_dTailPosFromSnap_cmm : DInt;
      TMP_xPlateIsInLimits : Bool;
      TMP_xPlateRespectControl : Bool;
      TMP_xXCutHeadDone : Bool;
      TMP_xXCutTailDone : Bool;
      TMP_dIndexCut : DInt;
      TMP_iValue : Int;
   END_VAR
   VAR CONSTANT
      CONST_DTHRDELPLATE_CMM : DInt := 700000;   // Threshold delete plate [mm/100]
      CONST_DTIMEOUTPLATEOFF_CMM : DInt := 200000;   // Timeout plate offset after a reset [mm/100]
      CONST_DSEARCH_HEAD : DInt := 1;   // Search only head limits
      CONST_DSEARCH_TAIL : DInt := 2;   // Search only tail limits
      CONST_DSEARCH_BOTH : DInt := 3;   // Search both head and tail
   END_VAR
   VAR_TEMP   // added for the SCL form of the ladder/FBD networks
      _w1 : Bool;
   END_VAR
BEGIN

REGION Network 1: Calculate OS of the general reset
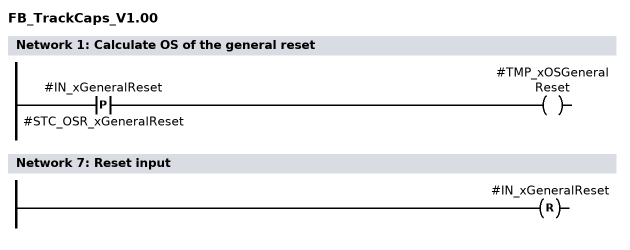
   RUNG wire#powerrail
      P_Contact(operand := #IN_xGeneralReset, bit := #STC_OSR_xGeneralReset)
      Coil( #TMP_xOSGeneralReset )
   END_RUNG
   // the same network as SCL:
   #_w1 := #IN_xGeneralReset AND NOT #STC_OSR_xGeneralReset;   // rising edge of #IN_xGeneralReset
   #STC_OSR_xGeneralReset := #IN_xGeneralReset;
   #TMP_xOSGeneralReset := #_w1;
END_REGION

REGION Network 2 (SCL): Reset tracking
   IF #TMP_xOSGeneralReset THEN

       #INO_tCaps.dLastInsertIndex := 0;
       #INO_tCaps.dTrackingHead := 0;
       #INO_tCaps.dTrackingTail := 0;
       #INO_tCaps.tLastPlacedCap := #INO_tCaps.tEmptyCap;
       #INO_tCaps.tNewCapToInsert := #INO_tCaps.tEmptyCap;
       #INO_tCaps.xInsertCapOnTrack := FALSE;
       #INO_tCaps.dLastTargetLineValue_cmm := #INO_tOptManager.tHMR.dLastOptLinePosition_cmm + #CONST_DTIMEOUTPLATEOFF_CMM; 
       #TMP_wValue := 0;

       SCATTER(IN:=#TMP_wValue,
           OUT=>#INO_tCaps.rgxNewCapAvailable);

       FOR #TMP_dIndex := 0 TO "DMAXTRACKCAP_IND" DO
           #INO_tCaps.rgtTrackCaps[#TMP_dIndex].dEncValueHeadSnaproll_cmm := 0;
           #INO_tCaps.rgtTrackCaps[#TMP_dIndex].dEncValueTailSnaproll_cmm := 0;
           #INO_tCaps.rgtTrackCaps[#TMP_dIndex].tCap := #INO_tCaps.tEmptyCap;
           #TMP_dwValue := 0;
           SCATTER(IN:= #TMP_dwValue, OUT=> #INO_tCaps.rgtTrackCaps[#TMP_dIndex].rgxMachineExecMask); 
       END_FOR;

       FOR #TMP_dIndex := 0 TO "DMAXTRACKMACHINE_IND" DO

           #INO_tCaps.rgtTrackMachine[#TMP_dIndex].tUserData.xGetPosReach := FALSE;
           #INO_tCaps.rgtTrackMachine[#TMP_dIndex].tAuxData.dActualMachineEncValue_cmm := 0;
           #INO_tCaps.rgtTrackMachine[#TMP_dIndex].tAuxData.dNextCapIndex := 0;
           #INO_tCaps.rgtTrackMachine[#TMP_dIndex].tAuxData.dPrevCapIndex := -1;
       END_FOR;
       //Update new cap to insert
       #INO_tCaps.tNewCapToInsert.dLength_cmm := 200000;
       #INO_tCaps.tNewCapToInsert.dWidth_cmm := 321000;
       #INO_tCaps.tNewCapToInsert.dThick_cmm := 500;
       #INO_tCaps.tNewCapToInsert.dFormat := 2;
       #INO_tCaps.tNewCapToInsert.dNumLites := 1;
       #INO_tCaps.tNewCapToInsert.dConvTotLength_cmm := 200000;
       #INO_tCaps.tNewCapToInsert.dGrossWidth_cmm := 330000;
       #INO_tCaps.tNewCapToInsert.dNetWidth_cmm := 330000;
       #INO_tCaps.tNewCapToInsert.rgtLites[0].dWidth_cmm := 321000;
       #INO_tCaps.tNewCapToInsert.rgtLites[0].dMainDestination := "DCULLETDESTMASK"; 

   END_IF;
END_REGION

REGION Network 3 (SCL): Insert plate on tracking
   IF #INO_tCaps.xInsertCapOnTrack THEN

       //Check if all the machines was informed about the new caps. If still mission to manage, exit.
       GATHER(IN:=#INO_tCaps.rgxNewCapAvailable,
              OUT=>#TMP_wValue);

      //RICORDARSI DI ATTIVARE QUESTO CONTROLLO 
      // IF #TMP_wValue <> 0 THEN
      //     RETURN;
      // END_IF;

       #TMP_dwValue := 16#FFFFFFFF;

       SCATTER(IN:=#TMP_dwValue,
               OUT=>#INO_tCaps.rgtTrackCaps[#INO_tCaps.dTrackingHead].rgxMachineExecMask);

       #INO_tCaps.rgtTrackCaps[#INO_tCaps.dTrackingHead].tCap := #INO_tCaps.tNewCapToInsert;
       #INO_tCaps.rgtTrackCaps[#INO_tCaps.dTrackingHead].dEncValueHeadSnaproll_cmm := #INO_tCaps.dLastTargetLineValue_cmm;
       #INO_tCaps.rgtTrackCaps[#INO_tCaps.dTrackingHead].dEncValueTailSnaproll_cmm := #INO_tCaps.dLastTargetLineValue_cmm + #INO_tCaps.tNewCapToInsert.dLength_cmm;
       #INO_tCaps.rgtTrackCaps[#INO_tCaps.dTrackingHead].tCap.dHeadPositionBTC := #INO_tCaps.dLastTargetLineValue_cmm;
       #INO_tCaps.rgtTrackCaps[#INO_tCaps.dTrackingHead].tCap.dTailPositionBTC := #INO_tCaps.dLastTargetLineValue_cmm + #INO_tCaps.tNewCapToInsert.dLength_cmm;

       #INO_tCaps.tNewCapToInsert.dHeadPositionBTC := #INO_tCaps.dLastTargetLineValue_cmm;
       #INO_tCaps.tNewCapToInsert.dTailPositionBTC := #INO_tCaps.dLastTargetLineValue_cmm + #INO_tCaps.tNewCapToInsert.dLength_cmm;
       #INO_tCaps.dLastTargetLineValue_cmm := #INO_tCaps.dLastTargetLineValue_cmm + #INO_tCaps.tNewCapToInsert.dLength_cmm;
       #INO_tCaps.dLastValidCapID := #INO_tCaps.tNewCapToInsert.rgtLites[#INO_tCaps.tNewCapToInsert.dNumLites-1].dID;
       #INO_tCaps.dNextValidCapID := #INO_tCaps.dLastValidCapID + 1;


       //Modification for ANCA to delete
       //#TMP_iValue := DWORD_TO_INT(#INO_tCaps.dNextValidCapID AND 16#0000FFFF);

       //IF #TMP_iValue < 0 THEN
       //    #INO_tCaps.dNextValidCapID := #INO_tCaps.dLastValidCapID + 32768;
       //END_IF;

       IF (#INO_tCaps.dNextValidCapID > "DMAXPLATEID") THEN

           #INO_tCaps.dNextValidCapID := 1;
           #INO_tCaps.dLastValidCapID := #INO_tCaps.dNextValidCapID;

       END_IF;

       //Send plate data for report
       #INO_tCaps.rgtTrackCaps[#INO_tCaps.dTrackingHead].tCap.tRequests.xUpdateDataBPSA := TRUE;     
       #INO_tCaps.rgtTrackCaps[#INO_tCaps.dTrackingHead].tCap.tRequests.xUpdateDataBPSB := TRUE;     

       #INO_tCaps.dLastInsertIndex := #INO_tCaps.dTrackingHead;

       IF (#INO_tCaps.dTrackingHead + 1) >= "DMAXTRACKCAP" THEN
           #INO_tCaps.dTrackingHead := 0;
       ELSE
           #INO_tCaps.dTrackingHead := #INO_tCaps.dTrackingHead + 1;
       END_IF;

       #INO_tCaps.tLastPlacedCap := #INO_tCaps.tNewCapToInsert;


       #TMP_wValue := 16#FFFF;

       SCATTER(IN:=#TMP_wValue,
               OUT=>#INO_tCaps.rgxNewCapAvailable);


       #INO_tCaps.xInsertCapOnTrack := FALSE;


   END_IF;
END_REGION

REGION Network 4 (SCL): Delete plate
   IF (#INO_tCaps.dTrackingHead <> #INO_tCaps.dTrackingTail) THEN

       #TMP_dValue_cmm := #INO_tEncoder.dActualEncoderCounter_cmm - #INO_tCaps.rgtTrackCaps[#INO_tCaps.dTrackingTail].dEncValueTailSnaproll_cmm;

       IF (#TMP_dValue_cmm > #CONST_DTHRDELPLATE_CMM) THEN

           #INO_tCaps.rgtTrackCaps[#INO_tCaps.dTrackingTail].dEncValueHeadSnaproll_cmm := 0;
           #INO_tCaps.rgtTrackCaps[#INO_tCaps.dTrackingTail].dEncValueTailSnaproll_cmm := 0;
           #INO_tCaps.rgtTrackCaps[#INO_tCaps.dTrackingTail].tCap := #INO_tCaps.tEmptyCap;
           #TMP_dwValue := 0;

           SCATTER(IN:= #TMP_dwValue, OUT=> #INO_tCaps.rgtTrackCaps[#INO_tCaps.dTrackingTail].rgxMachineExecMask); 

           IF (#INO_tCaps.dTrackingTail + 1) >= "DMAXTRACKCAP" THEN
               #INO_tCaps.dTrackingTail := 0;
           ELSE
               #INO_tCaps.dTrackingTail := #INO_tCaps.dTrackingTail + 1;
           END_IF;

       END_IF;

   END_IF;
END_REGION

REGION Network 5 (SCL): Machine checker
   FOR #TMP_dIndex := 0 TO "DMAXTRACKMACHINE_IND" DO

       //The machine last target line will be skipped because use a different count metod
       IF (#TMP_dIndex = "DMACHINEINDEX_LASTOPTLINE") THEN

           #TMP_dValue_cmm := #INO_tCaps.dLastTargetLineValue_cmm - #INO_tEncoder.dActualEncoderCounter_cmm;

           IF (#TMP_dValue_cmm <= #INO_tCaps.rgtTrackMachine["DMACHINEINDEX_LASTOPTLINE"].tUserData.dSetDistanceSnap_cmm) AND
               NOT (#INO_tCaps.rgtTrackMachine["DMACHINEINDEX_LASTOPTLINE"].tUserData.xGetPosReach) THEN

               #INO_tCaps.rgtTrackMachine["DMACHINEINDEX_LASTOPTLINE"].tUserData.dGetUpstremIndex := -1;
               #INO_tCaps.rgtTrackMachine["DMACHINEINDEX_LASTOPTLINE"].tUserData.dGetDownstreamIndex := -1;
               #INO_tCaps.rgtTrackMachine["DMACHINEINDEX_LASTOPTLINE"].tUserData.dGetEncValueOnSnap_cmm := #INO_tCaps.dLastTargetLineValue_cmm;
               #INO_tCaps.rgtTrackMachine["DMACHINEINDEX_LASTOPTLINE"].tUserData.xGetPosReach := TRUE;

           END_IF;

           CONTINUE;

       END_IF;

       //Calculate the actual encoder position of the machine
       #TMP_dActMachineEncValue_cmm := #INO_tEncoder.dActualEncoderCounter_cmm + 
                                       #INO_tCaps.rgtTrackMachine[#TMP_dIndex].tUserData.dSetDistanceSnap_cmm +
                                       REAL_TO_DINT(DINT_TO_REAL(#INO_tCaps.rgtTrackMachine[#TMP_dIndex].tUserData.dSetMachReacTime_ms) * #INO_tEncoder.rActSpeedValue_cmm_ms);

       //Next cap pointer
       #TMP_dIndexCap := #INO_tCaps.rgtTrackMachine[#TMP_dIndex].tAuxData.dNextCapIndex;

       //If plates are in the buffer
       IF (#INO_tCaps.dTrackingHead <> #INO_tCaps.dTrackingTail) THEN

           IF #INO_tCaps.rgtTrackCaps[#TMP_dIndexCap].rgxMachineExecMask[#TMP_dIndex] THEN

               #TMP_dValue_cmm := #TMP_dActMachineEncValue_cmm - #INO_tCaps.rgtTrackCaps[#TMP_dIndexCap].dEncValueHeadSnaproll_cmm;

               IF (#TMP_dValue_cmm >= 0) THEN

                   IF NOT (#INO_tCaps.rgtTrackMachine[#TMP_dIndex].tUserData.xGetPosReach) THEN

                       #INO_tCaps.rgtTrackMachine[#TMP_dIndex].tUserData.dGetUpstremIndex := #INO_tCaps.rgtTrackMachine[#TMP_dIndex].tAuxData.dNextCapIndex;
                       #INO_tCaps.rgtTrackMachine[#TMP_dIndex].tUserData.dGetDownstreamIndex := #INO_tCaps.rgtTrackMachine[#TMP_dIndex].tAuxData.dPrevCapIndex;
                       #INO_tCaps.rgtTrackMachine[#TMP_dIndex].tUserData.dGetEncValueOnSnap_cmm := #INO_tCaps.rgtTrackCaps[#TMP_dIndexCap].dEncValueHeadSnaproll_cmm;
                       #INO_tCaps.rgtTrackMachine[#TMP_dIndex].tUserData.xGetPosReach := TRUE;

                   END_IF;

                   #INO_tCaps.rgtTrackMachine[#TMP_dIndex].tAuxData.dPrevCapIndex := #INO_tCaps.rgtTrackMachine[#TMP_dIndex].tAuxData.dNextCapIndex;

                   IF (#INO_tCaps.rgtTrackMachine[#TMP_dIndex].tAuxData.dNextCapIndex + 1) >= "DMAXTRACKCAP" THEN
                       #INO_tCaps.rgtTrackMachine[#TMP_dIndex].tAuxData.dNextCapIndex := 0;
                   ELSE
                       #INO_tCaps.rgtTrackMachine[#TMP_dIndex].tAuxData.dNextCapIndex := #INO_tCaps.rgtTrackMachine[#TMP_dIndex].tAuxData.dNextCapIndex + 1;
                   END_IF;

                   #INO_tCaps.rgtTrackCaps[#TMP_dIndexCap].rgxMachineExecMask[#TMP_dIndex] := FALSE;

               END_IF;
           END_IF;
       END_IF;
   END_FOR;
END_REGION

REGION Network 6 (SCL): Search plates on tracking
   FOR #TMP_dIndex := 0 TO "DMAXELEMTRACKSEARCH_IND" DO

       IF #INO_tCaps.rgtTrackSearch[#TMP_dIndex].xRequestSearchPlate = TRUE AND 
           #INO_tCaps.rgtTrackSearch[#TMP_dIndex].xPlateFound = FALSE THEN

           //Request a tracking search. First aff all check the search condition. Search from the tail of the tracking until the head
           #TMP_dTail := #INO_tCaps.dTrackingTail;


           WHILE (#TMP_dTail <> #INO_tCaps.dTrackingHead) DO

               //Check if plate is present
               IF (#INO_tCaps.rgtTrackCaps[#TMP_dTail].tCap.dID <> 0) THEN

                   //Plate found calculate tail and head position from snaproll
                   #TMP_dHeadPosFromSnap_cmm := #INO_tCaps.rgtTrackCaps[#TMP_dTail].dEncValueHeadSnaproll_cmm - #INO_tEncoder.dActualEncoderCounter_cmm;
                   #TMP_dTailPosFromSnap_cmm := #INO_tCaps.rgtTrackCaps[#TMP_dTail].dEncValueTailSnaproll_cmm - #INO_tEncoder.dActualEncoderCounter_cmm;

                   //In according to the user request check if the plate is inside the limits requested
                   REGION PLATELIMITS

                   #TMP_xPlateIsInLimits := FALSE;

                   CASE #INO_tCaps.rgtTrackSearch[#TMP_dIndex].dSearchMode OF

                       #CONST_DSEARCH_HEAD:
                           IF #TMP_dHeadPosFromSnap_cmm >= #INO_tCaps.rgtTrackSearch[#TMP_dIndex].dMinHeadPosition_cmm AND
                               #TMP_dHeadPosFromSnap_cmm <= #INO_tCaps.rgtTrackSearch[#TMP_dIndex].dMaxHeadPosition_cmm THEN
                               #TMP_xPlateIsInLimits := TRUE;
                           END_IF;
                       #CONST_DSEARCH_TAIL:
                           IF #TMP_dTailPosFromSnap_cmm >= #INO_tCaps.rgtTrackSearch[#TMP_dIndex].dMinTailPosition_cmm AND
                               #TMP_dTailPosFromSnap_cmm <= #INO_tCaps.rgtTrackSearch[#TMP_dIndex].dMaxTailPosition_cmm THEN
                               #TMP_xPlateIsInLimits := TRUE;
                           END_IF;
                       #CONST_DSEARCH_BOTH: 
                           IF #TMP_dHeadPosFromSnap_cmm >= #INO_tCaps.rgtTrackSearch[#TMP_dIndex].dMinHeadPosition_cmm AND
                               #TMP_dHeadPosFromSnap_cmm <= #INO_tCaps.rgtTrackSearch[#TMP_dIndex].dMaxHeadPosition_cmm AND 
                               #TMP_dTailPosFromSnap_cmm >= #INO_tCaps.rgtTrackSearch[#TMP_dIndex].dMinTailPosition_cmm AND
                               #TMP_dTailPosFromSnap_cmm <= #INO_tCaps.rgtTrackSearch[#TMP_dIndex].dMaxTailPosition_cmm THEN
                               #TMP_xPlateIsInLimits := TRUE;
                           END_IF;
                   END_CASE;

                   END_REGION PLATELIMITS

                   //Plate in inside the limits, check the other control if are good
                   REGION CONTROLCHECK
                   #TMP_xPlateRespectControl := TRUE;

                   IF #TMP_xPlateIsInLimits THEN

                       IF #INO_tCaps.rgtTrackSearch[#TMP_dIndex].tSearchRequest.xLengthLessThan THEN

                           IF #INO_tCaps.rgtTrackCaps[#TMP_dTail].tCap.dLength_cmm >= #INO_tCaps.rgtTrackSearch[#TMP_dIndex].tSearchData.dLength_cmm THEN
                               #TMP_xPlateRespectControl := FALSE;
                           END_IF;

                       END_IF;

                       IF #INO_tCaps.rgtTrackSearch[#TMP_dIndex].tSearchRequest.xMainDestEqual THEN

                           IF #INO_tCaps.rgtTrackCaps[#TMP_dTail].tCap.rgtLites[0].dMainDestination <> #INO_tCaps.rgtTrackSearch[#TMP_dIndex].tSearchData.dMainDest_mask THEN
                               #TMP_xPlateRespectControl := FALSE;
                           END_IF;

                       END_IF;

                       IF #INO_tCaps.rgtTrackSearch[#TMP_dIndex].tSearchRequest.xCutDone THEN

                           #TMP_xXCutHeadDone := FALSE;
                           #TMP_xXCutTailDone := FALSE;

                           FOR #TMP_dIndexCut := 0 TO "DMAXXHEADS_IND" DO

                               IF #INO_tCaps.rgtTrackCaps[#TMP_dTail].tCap.tDone.rgxXCutDoneHead[#TMP_dIndexCut] THEN
                                   #TMP_xXCutHeadDone := TRUE;
                               END_IF;

                               IF #INO_tCaps.rgtTrackCaps[#TMP_dTail].tCap.tDone.rgxXCutDoneTail[#TMP_dIndexCut] THEN
                                   #TMP_xXCutTailDone := TRUE;
                               END_IF;

                           END_FOR;
                           IF NOT #TMP_xXCutHeadDone OR NOT #TMP_xXCutTailDone THEN
                               #TMP_xPlateRespectControl := FALSE;
                           END_IF;

                       END_IF;

                       //The plate is valid. Compile the output data   
                       IF #TMP_xPlateRespectControl THEN
                           #INO_tCaps.rgtTrackSearch[#TMP_dIndex].dFoundTrackIndex := #TMP_dTail;                 
                           #INO_tCaps.rgtTrackSearch[#TMP_dIndex].xPlateFound := TRUE;
                           //Exit the while cycle. The search is terminated
                           EXIT;
                       END_IF;
                   END_IF;
                   END_REGION CONTROLCHECK

               END_IF;

               //Increment the tail
               IF (#TMP_dTail + 1) >= "DMAXTRACKCAP" THEN
                   #TMP_dTail := 0;
               ELSE
                   #TMP_dTail+= 1;
               END_IF;

           END_WHILE;
           //Move the validation ID 
           #INO_tCaps.rgtTrackSearch[#TMP_dIndex].dAnalyzedID := #INO_tCaps.rgtTrackSearch[#TMP_dIndex].dRequestID;
       END_IF;

   END_FOR;
END_REGION

REGION Network 7: Reset input
   RUNG wire#powerrail
      R_Coil( #IN_xGeneralReset )
   END_RUNG
   // the same network as SCL:
   #IN_xGeneralReset := FALSE;
END_REGION
END_FUNCTION_BLOCK

// folder: 03_Programs_Logics/MCC1200/03_CrossCut

